'~S001R16 EE (Clmp Not Clsd, Slide Not Advd, Pin Not Retd, Still Opn, Still Ret) S001R16B#.O.A S001R16B#.I.## FB2[234].16'; 7505 '~S001R16 EE (Clmp Not Opnd, Slide Not Retd, Pin Not Advd, Still Clsd, Still Adv) S001R16B#.O.A S001R16B#.I.## FB2[234].17'; 7506 '~S001R16 EE (Clmp Not Clsd, Slide Not Advd, Pin Not Retd, Still Opn, Still Ret) S001R16B#.O.A S001R16B#.I.## FB2[234].18'; 7507 '~S001R16 EE (Clmp Not Opnd, Slide Not Retd, Pin Not Advd, Still Clsd, Still Adv) S001R16B#.O.A S001R16B#.I.## FB2[234].19'; 7508 '~S001R16 EE (Clmp Not Clsd, Slide Not Advd, Pin Not Retd, Still Opn, Still Ret) S001R16B#.O.A S001R16B#.I.## FB2[234].20'; 7509 '~S001R16 EE (Clmp Not Opnd, Slide Not Retd, Pin Not Advd, Still Clsd, Still Adv) S001R16B#.O.A S001R16B#.I.## FB2[234].21'; 7510 '~S001R16 EE (Clmp Not Clsd, Slide Not Advd, Pin Not Retd, Still Opn, Still Ret) S001R16B#.O.A S001R16B#.I.## FB2[234].22'; 7511 '~S001R16 EE (Clmp Not Opnd, Slide Not Retd, Pin Not Advd, Still Clsd, Still Adv) S001R16B#.O.A S001R16B#.I.## FB2[234].23'; 7512 '~S001R16 EE (Clmp Not Clsd, Slide Not Advd, Pin Not Retd, Still Opn, Still Ret) S001R16B#.O.A S001R16B#.I.## FB2[234].24'; 7513 '~S001R16 EE (Clmp Not Opnd, Slide Not Retd, Pin Not Advd, Still Clsd, Still Adv) S001R16B#.O.A S001R16B#.I.## FB2[234].25'; 7514 '~S001R16 EE (Clmp Not Clsd, Slide Not Advd, Pin Not Retd, Still Opn, Still Ret) S001R16B#.O.A S001R16B#.I.## FB2[234].26'; 7515 '~S001R16 EE (Clmp Not Opnd, Slide Not Retd, Pin Not Advd, Still Clsd, Still Adv) S001R16B#.O.A S001R16B#.I.## FB2[234].27'; 7516 '~S001R16 EE (Clmp Not Clsd, Slide Not Advd, Pin Not Retd, Still Opn, Still Ret) S001R16B#.O.A S001R16B#.I.## FB2[234].28'; 7517 '~S001R16 EE (Clmp Not Opnd, Slide Not Retd, Pin Not Advd, Still Clsd, Still Adv) S001R16B#.O.A S001R16B#.I.## FB2[234].29'; 7518 '~S001R16 EE (Clmp Not Clsd, Slide Not Advd, Pin Not Retd, Still Opn, Still Ret) S001R16B#.O.A S001R16B#.I.## FB2[234].30'; 7519 '~S001R16 EE (Clmp Not Opnd, Slide Not Retd, Pin Not Advd, Still Clsd, Still Adv) S001R16B#.O.A S001R16B#.I.## FB2[234].31'; 7520 '~S001R16 EE (Clmp Not Clsd, Slide Not Advd, Pin Not Retd, Still Opn, Still Ret) S001R16B#.O.A S001R16B#.I.## FB2[235].0'; 7521 '~S001R16 EE (Clmp Not Opnd, Slide Not Retd, Pin Not Advd, Still Clsd, Still Adv) S001R16B#.O.A S001R16B#.I.## FB2[235].1'; 7522 '~S001R16 EE (Clmp Not Clsd, Slide Not Advd, Pin Not Retd, Still Opn, Still Ret) S001R16B#.O.A S001R16B#.I.## FB2[235].2'; 7523 '~S001R16 EE (Clmp Not Opnd, Slide Not Retd, Pin Not Advd, Still Clsd, Still Adv) S001R16B#.O.A S001R16B#.I.## FB2[235].3'; 7524 '~S001R16 EE (Clmp Not Clsd, Slide Not Advd, Pin Not Retd, Still Opn, Still Ret) S001R16B#.O.A S001R16B#.I.## FB2[235].4'; 7525 '~S001R16 EE (Clmp Not Opnd, Slide Not Retd, Pin Not Advd, Still Clsd, Still Adv) S001R16B#.O.A S001R16B#.I.## FB2[235].5'; 7526 '~S001R16 EE (Clmp Not Clsd, Slide Not Advd, Pin Not Retd, Still Opn, Still Ret) S001R16B#.O.A S001R16B#.I.## FB2[235].6'; 7527 '~S001R16 EE (Clmp Not Opnd, Slide Not Retd, Pin Not Advd, Still Clsd, Still Adv) S001R16B#.O.A S001R16B#.I.## FB2[235].7'; 7528 '~S001R16 EE (Clmp Not Clsd, Slide Not Advd, Pin Not Retd, Still Opn, Still Ret) S001R16B#.O.A S001R16B#.I.## FB2[235].8'; 7529 '~S001R16 EE (Clmp Not Opnd, Slide Not Retd, Pin Not Advd, Still Clsd, Still Adv) S001R16B#.O.A S001R16B#.I.## FB2[235].9'; 7530 '~S001R16 EE (Clmp Not Clsd, Slide Not Advd, Pin Not Retd, Still Opn, Still Ret) S001R16B#.O.A S001R16B#.I.## FB2[235].10'; 7531 '~S001R16 EE (Clmp Not Opnd, Slide Not Retd, Pin Not Advd, Still Clsd, Still Adv) S001R16B#.O.A S001R16B#.I.## FB2[235].11'; 7532 '~S001R16 EE (Clmp Not Clsd, Slide Not Advd, Pin Not Retd, Still Opn, Still Ret) S001R16B#.O.A S001R16B#.I.## FB2[235].12'; 7533 '~S001R16 EE (Clmp Not Opnd, Slide Not Retd, Pin Not Advd, Still Clsd, Still Adv) S001R16B#.O.A S001R16B#.I.## FB2[235].13'; 7534 '~S001R16 EE (Clmp Not Clsd, Slide Not Advd, Pin Not Retd, Still Opn, Still Ret) S001R16B#.O.A S001R16B#.I.## FB2[235].14'; 7535 '~S001R16 EE (Clmp Not Opnd, Slide Not Retd, Pin Not Advd, Still Clsd, Still Adv) S001R16B#.O.A S001R16B#.I.## FB2[235].15'; 7536 '~S001R16 EE (Clmp Not Clsd, Slide Not Advd, Pin Not Retd, Still Opn, Still Ret) S001R16B#.O.A S001R16B#.I.## FB2[235].16'; 7537 '~S001R16 EE (Clmp Not Opnd, Slide Not Retd, Pin Not Advd, Still Clsd, Still Adv) S001R16B#.O.A S001R16B#.I.## FB2[235].17'; 7538 '~S001R16 EE (Clmp Not Clsd, Slide Not Advd, Pin Not Retd, Still Opn, Still Ret) S001R16B#.O.A S001R16B#.I.## FB2[235].18'; 7539 '~S001R16 EE (Clmp Not Opnd, Slide Not Retd, Pin Not Advd, Still Clsd, Still Adv) S001R16B#.O.A S001R16B#.I.## FB2[235].19'; 7540 '~S001R16 EE (Clmp Not Clsd, Slide Not Advd, Pin Not Retd, Still Opn, Still Ret) S001R16B#.O.A S001R16B#.I.## FB2[235].20'; 7541 '~S001R16 EE (Clmp Not Opnd, Slide Not Retd, Pin Not Advd, Still Clsd, Still Adv) S001R16B#.O.A S001R16B#.I.## FB2[235].21'; 7542 '~S001R16 EE (Clmp Not Clsd, Slide Not Advd, Pin Not Retd, Still Opn, Still Ret) S001R16B#.O.A S001R16B#.I.## FB2[235].22'; 7543 '~S001R16 EE (Clmp Not Opnd, Slide Not Retd, Pin Not Advd, Still Clsd, Still Adv) S001R16B#.O.A S001R16B#.I.## FB2[235].23'; 7544 '~S001R16 EE (Clmp Not Clsd, Slide Not Advd, Pin Not Retd, Still Opn, Still Ret) S001R16B#.O.A S001R16B#.I.## FB2[235].24'; 7545 '~S001R16 EE (Clmp Not Opnd, Slide Not Retd, Pin Not Advd, Still Clsd, Still Adv) S001R16B#.O.A S001R16B#.I.## FB2[235].25'; 7546 '~S001R16 EE (Clmp Not Clsd, Slide Not Advd, Pin Not Retd, Still Opn, Still Ret) S001R16B#.O.A S001R16B#.I.## FB2[235].26'; 7547 '~S001R16 EE (Clmp Not Opnd, Slide Not Retd, Pin Not Advd, Still Clsd, Still Adv) S001R16B#.O.A S001R16B#.I.## FB2[235].27'; 7548 '~S001R16 EE (Clmp Not Clsd, Slide Not Advd, Pin Not Retd, Still Opn, Still Ret) S001R16B#.O.A S001R16B#.I.## FB2[235].28'; 7549 '~S001R16 EE (Clmp Not Opnd, Slide Not Retd, Pin Not Advd, Still Clsd, Still Adv) S001R16B#.O.A S001R16B#.I.## FB2[235].29'; 7550 '~S001R16 EE (Clmp Not Clsd, Slide Not Advd, Pin Not Retd, Still Opn, Still Ret) S001R16B#.O.A S001R16B#.I.## FB2[235].30'; 7551 '~S001R16 EE (Clmp Not Opnd, Slide Not Retd, Pin Not Advd, Still Clsd, Still Adv) S001R16B#.O.A S001R16B#.I.## FB2[235].31'; 7552 '~Spare FB2[236].0'; 7553 '~Spare FB2[236].1'; 7554 '~Spare FB2[236].2'; 7555 '~Spare FB2[236].3'; 7556 '~Spare FB2[236].4'; 7557 '~Spare FB2[236].5'; 7558 '~Spare FB2[236].6'; 7559 '~Spare FB2[236].7'; 7560 '~Spare FB2[236].8'; 7561 '~Spare FB2[236].9'; 7562 '~Spare FB2[236].10'; 7563 '~Spare FB2[236].11'; 7564 '~Spare FB2[236].12'; 7565 '~Spare FB2[236].13'; 7566 '~Spare FB2[236].14'; 7567 '~Spare FB2[236].15'; 7568 '~Spare FB2[236].16'; 7569 '~Spare FB2[236].17'; 7570 '~Spare FB2[236].18'; 7571 '~Spare FB2[236].19'; 7572 '~Spare FB2[236].20'; 7573 '~Spare FB2[236].21'; 7574 '~Spare FB2[236].22'; 7575 '~Spare FB2[236].23'; 7576 '~Spare FB2[236].24'; 7577 '~Spare FB2[236].25'; 7578 '~Spare FB2[236].26'; 7579 '~Spare FB2[236].27'; 7580 '~Spare FB2[236].28'; 7581 '~Spare FB2[236].29'; 7582 '~Spare FB2[236].30'; 7583 '~Spare FB2[236].31'; 7584 '~Spare FB2[237].0'; 7585 '~Spare FB2[237].1'; 7586 '~Spare FB2[237].2'; 7587 '~Spare FB2[237].3'; 7588 '~Spare FB2[237].4'; 7589 '~Spare FB2[237].5'; 7590 '~Spare FB2[237].6'; 7591 '~Spare FB2[237].7'; 7592 '~Spare FB2[237].8'; 7593 '~Spare FB2[237].9'; 7594 '~Spare FB2[237].10'; 7595 '~Spare FB2[237].11'; 7596 '~Spare FB2[237].12'; 7597 '~Spare FB2[237].13'; 7598 '~Spare FB2[237].14'; 7599 '~Spare FB2[237].15'; 7600 '~Spare FB2[237].16'; 7601 '~Spare FB2[237].17'; 7602 '~Spare FB2[237].18'; 7603 '~Spare FB2[237].19'; 7604 '~Spare FB2[237].20'; 7605 '~Spare FB2[237].21'; 7606 '~Spare FB2[237].22'; 7607 '~Spare FB2[237].23'; 7608 '~Spare FB2[237].24'; 7609 '~Spare FB2[237].25'; 7610 '~Spare FB2[237].26'; 7611 '~Spare FB2[237].27'; 7612 '~Spare FB2[237].28'; 7613 '~Spare FB2[237].29'; 7614 '~Spare FB2[237].30'; 7615 '~Spare FB2[237].31'; 7616 '~Spare FB2[238].0'; 7617 '~Spare FB2[238].1'; 7618 '~Spare FB2[238].2'; 7619 '~Spare FB2[238].3'; 7620 '~Spare FB2[238].4'; 7621 '~Spare FB2[238].5'; 7622 '~Spare FB2[238].6'; 7623 '~Spare FB2[238].7'; 7624 '~Spare FB2[238].8'; 7625 '~Spare FB2[238].9'; 7626 '~Spare FB2[238].10'; 7627 '~Spare FB2[238].11'; 7628 '~Spare FB2[238].12'; 7629 '~Spare FB2[238].13'; 7630 '~Spare FB2[238].14'; 7631 '~Spare FB2[238].15'; 7632 '~Spare FB2[238].16'; 7633 '~Spare FB2[238].17'; 7634 '~Spare FB2[238].18'; 7635 '~Spare FB2[238].19'; 7636 '~Spare FB2[238].20'; 7637 '~Spare FB2[238].21'; 7638 '~Spare FB2[238].22'; 7639 '~Spare FB2[238].23'; 7640 '~Spare FB2[238].24'; 7641 '~Spare FB2[238].25'; 7642 '~Spare FB2[238].26'; 7643 '~Spare FB2[238].27'; 7644 '~Spare FB2[238].28'; 7645 '~Spare FB2[238].29'; 7646 '~Spare FB2[238].30'; 7647 '~Spare FB2[238].31'; 7648 '~S001R16 (Peripheral Tool 1) Vlv/Otpt 1 Failed S001R16F#B#.O.# (Cls Clmps, Adv Slide, Ret Pins) FB2[239].0'; 7649 '~S001R16 (Peripheral Tool 1) Vlv/Otpt 1 Failed S001R16F#B#.O.# (Opn Clmps, Ret Slide, Adv Pins) FB2[239].1'; 7650 '~S001R16 (Peripheral Tool 1) Vlv/Otpt 2 Failed S001R16F#B#.O.# (Cls Clmps, Adv Slide, Ret Pins) FB2[239].2'; 7651 '~S001R16 (Peripheral Tool 1) Vlv/Otpt 2 Failed S001R16F#B#.O.# (Opn Clmps, Ret Slide, Adv Pins) FB2[239].3'; 7652 '~S001R16 (Peripheral Tool 1) Vlv/Otpt 3 Failed S001R16F#B#.O.# (Cls Clmps, Adv Slide, Ret Pins) FB2[239].4'; 7653 '~S001R16 (Peripheral Tool 1) Vlv/Otpt 3 Failed S001R16F#B#.O.# (Opn Clmps, Ret Slide, Adv Pins) FB2[239].5'; 7654 '~S001R16 (Peripheral Tool 1) Vlv/Otpt 4 Failed S001R16F#B#.O.# (Cls Clmps, Adv Slide, Ret Pins) FB2[239].6'; 7655 '~S001R16 (Peripheral Tool 1) Vlv/Otpt 4 Failed S001R16F#B#.O.# (Opn Clmps, Ret Slide, Adv Pins) FB2[239].7'; 7656 '~U-#### (Clmp Not Clsd, Slide Not Advd, Pin Not Retd, Still Opnd, Still Retd) S001R16F#.B#.O.# FB2[239].8'; 7657 '~U-#### (Clmp Not Opnd, Slide Not Retd, Pin Not Advd, Still Clsd, Still Advd) S001R16F#.B#.O.# FB2[239].9'; 7658 '~U-#### (Clmp Not Clsd, Slide Not Advd, Pin Not Retd, Still Opnd, Still Retd) S001R16F#.B#.O.# FB2[239].10'; 7659 '~U-#### (Clmp Not Opnd, Slide Not Retd, Pin Not Advd, Still Clsd, Still Advd) S001R16F#.B#.O.# FB2[239].11'; 7660 '~U-#### (Clmp Not Clsd, Slide Not Advd, Pin Not Retd, Still Opnd, Still Retd) S001R16F#.B#.O.# FB2[239].12'; 7661 '~U-#### (Clmp Not Opnd, Slide Not Retd, Pin Not Advd, Still Clsd, Still Advd) S001R16F#.B#.O.# FB2[239].13'; 7662 '~U-#### (Clmp Not Clsd, Slide Not Advd, Pin Not Retd, Still Opnd, Still Retd) S001R16F#.B#.O.# FB2[239].14'; 7663 '~U-#### (Clmp Not Opnd, Slide Not Retd, Pin Not Advd, Still Clsd, Still Advd) S001R16F#.B#.O.# FB2[239].15'; 7664 '~S001R16 (Peripheral Tool 2) Vlv/Otpt 1 Failed S001R16F#B#.O.# (Cls Clmps, Adv Slide, Ret Pins) FB2[239].16'; 7665 '~S001R16 (Peripheral Tool 2) Vlv/Otpt 1 Failed S001R16F#B#.O.# (Opn Clmps, Ret Slide, Adv Pins) FB2[239].17'; 7666 '~S001R16 (Peripheral Tool 2) Vlv/Otpt 2 Failed S001R16F#B#.O.# (Cls Clmps, Adv Slide, Ret Pins) FB2[239].18'; 7667 '~S001R16 (Peripheral Tool 2) Vlv/Otpt 2 Failed S001R16F#B#.O.# (Opn Clmps, Ret Slide, Adv Pins) FB2[239].19'; 7668 '~S001R16 (Peripheral Tool 2) Vlv/Otpt 3 Failed S001R16F#B#.O.# (Cls Clmps, Adv Slide, Ret Pins) FB2[239].20'; 7669 '~S001R16 (Peripheral Tool 2) Vlv/Otpt 3 Failed S001R16F#B#.O.# (Opn Clmps, Ret Slide, Adv Pins) FB2[239].21'; 7670 '~S001R16 (Peripheral Tool 2) Vlv/Otpt 4 Failed S001R16F#B#.O.# (Cls Clmps, Adv Slide, Ret Pins) FB2[239].22'; 7671 '~S001R16 (Peripheral Tool 2) Vlv/Otpt 4 Failed S001R16F#B#.O.# (Opn Clmps, Ret Slide, Adv Pins) FB2[239].23'; 7672 '~U-#### (Clmp Not Clsd, Slide Not Advd, Pin Not Retd, Still Opnd, Still Retd) S001R16F#.B#.O.# FB2[239].24'; 7673 '~U-#### (Clmp Not Opnd, Slide Not Retd, Pin Not Advd, Still Clsd, Still Advd) S001R16F#.B#.O.# FB2[239].25'; 7674 '~U-#### (Clmp Not Clsd, Slide Not Advd, Pin Not Retd, Still Opnd, Still Retd) S001R16F#.B#.O.# FB2[239].26'; 7675 '~U-#### (Clmp Not Opnd, Slide Not Retd, Pin Not Advd, Still Clsd, Still Advd) S001R16F#.B#.O.# FB2[239].27'; 7676 '~U-#### (Clmp Not Clsd, Slide Not Advd, Pin Not Retd, Still Opnd, Still Retd) S001R16F#.B#.O.# FB2[239].28'; 7677 '~U-#### (Clmp Not Opnd, Slide Not Retd, Pin Not Advd, Still Clsd, Still Advd) S001R16F#.B#.O.# FB2[239].29'; 7678 '~U-#### (Clmp Not Clsd, Slide Not Advd, Pin Not Retd, Still Opnd, Still Retd) S001R16F#.B#.O.# FB2[239].30'; 7679 '~U-#### (Clmp Not Opnd, Slide Not Retd, Pin Not Advd, Still Clsd, Still Advd) S001R16F#.B#.O.# FB2[239].31'; 7680 '~Spare FB2[240].0'; 7681 '~Spare FB2[240].1'; 7682 '~Spare FB2[240].2'; 7683 '~Spare FB2[240].3'; 7684 '~Spare FB2[240].4'; 7685 '~Spare FB2[240].5'; 7686 '~Spare FB2[240].6'; 7687 '~Spare FB2[240].7'; 7688 '~Spare FB2[240].8'; 7689 '~Spare FB2[240].9'; 7690 '~Spare FB2[240].10'; 7691 '~Spare FB2[240].11'; 7692 '~Spare FB2[240].12'; 7693 '~Spare FB2[240].13'; 7694 '~Spare FB2[240].14'; 7695 '~Spare FB2[240].15'; 7696 '~Spare FB2[240].16'; 7697 '~Spare FB2[240].17'; 7698 '~Spare FB2[240].18'; 7699 '~Spare FB2[240].19'; 7700 '~Spare FB2[240].20'; 7701 '~Spare FB2[240].21'; 7702 '~Spare FB2[240].22'; 7703 '~Spare FB2[240].23'; 7704 '~Spare FB2[240].24'; 7705 '~Spare FB2[240].25'; 7706 '~Spare FB2[240].26'; 7707 '~Spare FB2[240].27'; 7708 '~Spare FB2[240].28'; 7709 '~Spare FB2[240].29'; 7710 '~Spare FB2[240].30'; 7711 '~Spare FB2[240].31'; 7712 '~Spare FB2[241].0'; 7713 '~Spare FB2[241].1'; 7714 '~Spare FB2[241].2'; 7715 '~Spare FB2[241].3'; 7716 '~Spare FB2[241].4'; 7717 '~Spare FB2[241].5'; 7718 '~Spare FB2[241].6'; 7719 '~Spare FB2[241].7'; 7720 '~Spare FB2[241].8'; 7721 '~Spare FB2[241].9'; 7722 '~Spare FB2[241].10'; 7723 '~Spare FB2[241].11'; 7724 '~Spare FB2[241].12'; 7725 '~Spare FB2[241].13'; 7726 '~Spare FB2[241].14'; 7727 '~Spare FB2[241].15'; 7728 '~Spare FB2[241].16'; 7729 '~Spare FB2[241].17'; 7730 '~Spare FB2[241].18'; 7731 '~Spare FB2[241].19'; 7732 '~Spare FB2[241].20'; 7733 '~Spare FB2[241].21'; 7734 '~Spare FB2[241].22'; 7735 '~Spare FB2[241].23'; 7736 '~Spare FB2[241].24'; 7737 '~Spare FB2[241].25'; 7738 '~Spare FB2[241].26'; 7739 '~Spare FB2[241].27'; 7740 '~Spare FB2[241].28'; 7741 '~Spare FB2[241].29'; 7742 '~Spare FB2[241].30'; 7743 '~Spare FB2[241].31'; 7744 '~Spare FB2[242].0'; 7745 '~Spare FB2[242].1'; 7746 '~Spare FB2[242].2'; 7747 '~Spare FB2[242].3'; 7748 '~Spare FB2[242].4'; 7749 '~Spare FB2[242].5'; 7750 '~Spare FB2[242].6'; 7751 '~Spare FB2[242].7'; 7752 '~Spare FB2[242].8'; 7753 '~Spare FB2[242].9'; 7754 '~Spare FB2[242].10'; 7755 '~Spare FB2[242].11'; 7756 '~Spare FB2[242].12'; 7757 '~Spare FB2[242].13'; 7758 '~Spare FB2[242].14'; 7759 '~Spare FB2[242].15'; 7760 '~Spare FB2[242].16'; 7761 '~Spare FB2[242].17'; 7762 '~Spare FB2[242].18'; 7763 '~Spare FB2[242].19'; 7764 '~Spare FB2[242].20'; 7765 '~Spare FB2[242].21'; 7766 '~Spare FB2[242].22'; 7767 '~Spare FB2[242].23'; 7768 '~Spare FB2[242].24'; 7769 '~Spare FB2[242].25'; 7770 '~Spare FB2[242].26'; 7771 '~Spare FB2[242].27'; 7772 '~Spare FB2[242].28'; 7773 '~Spare FB2[242].29'; 7774 '~Spare FB2[242].30'; 7775 '~Spare FB2[242].31'; 7776 '~Spare FB2[243].0'; 7777 '~Spare FB2[243].1'; 7778 '~Spare FB2[243].2'; 7779 '~Spare FB2[243].3'; 7780 '~Spare FB2[243].4'; 7781 '~Spare FB2[243].5'; 7782 '~Spare FB2[243].6'; 7783 '~Spare FB2[243].7'; 7784 '~Spare FB2[243].8'; 7785 '~Spare FB2[243].9'; 7786 '~Spare FB2[243].10'; 7787 '~Spare FB2[243].11'; 7788 '~Spare FB2[243].12'; 7789 '~Spare FB2[243].13'; 7790 '~Spare FB2[243].14'; 7791 '~Spare FB2[243].15'; 7792 '~Spare FB2[243].16'; 7793 '~Spare FB2[243].17'; 7794 '~Spare FB2[243].18'; 7795 '~Spare FB2[243].19'; 7796 '~Spare FB2[243].20'; 7797 '~Spare FB2[243].21'; 7798 '~Spare FB2[243].22'; 7799 '~Spare FB2[243].23'; 7800 '~Spare FB2[243].24'; 7801 '~Spare FB2[243].25'; 7802 '~Spare FB2[243].26'; 7803 '~Spare FB2[243].27'; 7804 '~Spare FB2[243].28'; 7805 '~Spare FB2[243].29'; 7806 '~Spare FB2[243].30'; 7807 '~Spare FB2[243].31'; 7808 '~S001R09CN.I.RbtCtrlFlt - Control Fault FB2[244].0'; 7809 '~S001R09CN.I.CollDetect - Collision Detect FB2[244].1'; 7810 '~S001R09CN.Ix.RbtPromptBox - View Prompt Box at Teach Pendant FB2[244].2'; 7811 '~Spare FB2[244].3'; 7812 '~Spare FB2[244].4'; 7813 '~Spare FB2[244].5'; 7814 '~Spare FB2[244].6'; 7815 '~Spare FB2[244].7'; 7816 '~Spare FB2[244].8'; 7817 '~Spare FB2[244].9'; 7818 '~Spare FB2[244].10'; 7819 '~S001R09CN.I.Wc1WldFlt -Weld Controller 1 Weld Fault FB2[244].11'; 7820 '~S001R09CN.I.Wc1Flt - Weld Timer Flt - Depress Man Weld To Continue FB2[244].12'; 7821 '~S001R09CN.I.Wc1SGunFlt - Weld Controller 1 Servo Gun Fault FB2[244].13'; 7822 '~S001R09CN.I.Wc1SGunMtrTempFlt - Cntrl 1 Servo Gun Motor Over Temp FB2[244].14'; 7823 '~S001R09CN.I.Td1MtrFlt - Tip Dress 1 Motor Fault FB2[244].15'; 7824 '~S001R09CN.I.WC1XfmrTempFlt - Weld Cntrl 1 Transformer Over Temp FB2[244].16'; 7825 '~S001R09CN.I.AutoTipChng1Flt - Auto Tip Changer 1 Fault FB2[244].17'; 7826 '~S001R09CN.I.Slr1NotReady - Seal Controller 1 Not Ready FB2[244].18'; 7827 '~S001R09CN.I.Slr1MajorFlt - Seal Controller 1 Major Fault FB2[244].19'; 7828 '~S001R09CN.I.Slr1VolNotOk - Seal Controller 1 Volume Not Ok Fault FB2[244].20'; 7829 '~S001R09CN.I.Slr1PurgeFlt - Seal Controller 1 Purge Fault FB2[244].21'; 7830 '~S001R09CN.I.Slr1DoserNot Filled - Seal Cntrl 1 Doser Not Filled FB2[244].22'; 7831 '~S001R09CN.I.Slr1No2ClnMxr - Seal Cntrl1 No 2C In Mixer Fault FB2[244].23'; 7832 '~S001R09CN.I.Slr1NzlBroken - Seal Controller 1 Nozzle Broken Fault FB2[244].24'; 7833 '~S001R09CN.I.Slr1NozzleChgReq - Seal Cntrl1 Nozzle Change Reqd FB2[244].25'; 7834 '~S001R09CN.I.Slr1CycleInterrupted - Seal Cntrl1 Cycle Interrupted FB2[244].26'; 7835 '~S001R09CN.I.Stdw1Flt - Stud Weld 1 Weld Fault FB2[244].27'; 7836 '~S001R09CN.I.Stdw1DlyExcdd - Stud Weld 1 Time Delay Exceeded Flt FB2[244].28'; 7837 '~S001R09CN.I.Stdw1Maint Reqd - Stud Weld 1 Maintenance Required FB2[244].29'; 7838 '~S001R09CN.I.Stdw1Reject - Stud Weld 1 art Reject Fault FB2[244].30'; 7839 '~S001R09CN.I.Rvt1Flt - Rivet Controller 1 Fault FB2[244].31'; 7840 '~S001R09CN.I.Rvt1DlyExcdd - Rivet Cntrl 1 Time Delay Exceeded Flt FB2[245].0'; 7841 '~S001R09CN.I.AutoPulledTipByp1 - Auto Pulled Tip Bypass 1 FB2[245].1'; 7842 '~S001R09CN.I.StdWld1EquipmentFlt - Stud Weld 1 Equipment Fault FB2[245].2'; 7843 '~S001R09CN.I.StdWld1BrcktNotPresent - Stud Weld 1 Bracket Not Pres FB2[245].3'; 7844 '~S001R09CN.I.PierceFlt - Pierce Fault FB2[245].4'; 7845 '~S001R09CN.I.NoVisionMeasErr - Vision System Measurement Error FB2[245].5'; 7846 '~S001R09CN.I.VisionSysCalErr - Vision System Calibration Fault FB2[245].6'; 7847 '~S001R09CN.I.VisionSysErr - Vision System Error FB2[245].7'; 7848 '~S001R09CN.I.RackOutOfTolerance - Vision Sys Rack Out Of Tolerance FB2[245].8'; 7849 '~S001R09CN.Ix.TorqFlt - Torque Not Ok FB2[245].9'; 7850 '~S001R09CN.Ix.MwFlt - Mig Weld Controller Fault FB2[245].10'; 7851 '~S001R09CN.Ix.MwWireStuckFlt - Mig Welder Wire Stuck FB2[245].11'; 7852 '~S001R09CN.Ix.MwWldFlt - Mig Welder Bad Bronze Weld Indicator Flt FB2[245].12'; 7853 '~S001R09CN.I.O.TipChngReqd1 - Weld Cntrl 1 Tip Change Required FB2[245].13'; 7854 '~S001R09CN.I.M.NutDetectFlt1 - Nut Welder 1 Nut Detection Fault FB2[245].14'; 7855 '~S001R09CN.I.M.NutProjFlt1 - Nut Welder 1 Weld Not In Tolerance FB2[245].15'; 7856 '~S001R09CN.M.WrongRivetAtNose - Remove Wrong Rivet At Nose FB2[245].16'; 7857 '~S001R09CN.Ix.MwWldLimitErr - Mig Welder CurrentVoltage Out of Tolerance FB2[245].17'; 7858 '~S001R09CN.Ix.MigRdy Mig Welder Not Ready FB2[245].18'; 7859 '~Spare FB2[245].19'; 7860 '~Spare FB2[245].20'; 7861 '~S001R09CN.I.Wc2WldFlt -Weld Controller 2 Weld Fault FB2[245].21'; 7862 '~S001R09CN.I.Wc2Flt - Weld Timer Flt - Depress Man Weld To Continue FB2[245].22'; 7863 '~S001R09CN.I.Wc2SGunFlt - Weld Controller 2 Servo Gun Fault FB2[245].23'; 7864 '~S001R09CN.I.Wc2SGunMtrTempFlt - Cntrl 2 Servo Gun Motor Over Temp FB2[245].24'; 7865 '~S001R09CN.I.Td2MtrFlt - Tip Dress 2 Motor Fault FB2[245].25'; 7866 '~S001R09CN.I.WC2XfmrTempFlt - Weld Cntrl 2 Transformer Over Temp FB2[245].26'; 7867 '~S001R09CN.I.AutoTipChng2Flt - Auto Tip Changer 2 Fault FB2[245].27'; 7868 '~S001R09CN.I.Slr2NotReady - Seal Controller 2 Not Ready FB2[245].28'; 7869 '~S001R09CN.I.Slr2MajorFlt - Seal Controller 2 Major Fault FB2[245].29'; 7870 '~S001R09CN.I.Slr2VolNotOk - Seal Controller 2 Volume Not Ok Fault FB2[245].30'; 7871 '~S001R09CN.I.Slr2PurgeFlt - Seal Controller 2 Purge Fault FB2[245].31'; 7872 '~S001R09CN.I.Slr2DoserNot Filled - Seal Cntrl 2 Doser Not Filled FB2[246].0'; 7873 '~S001R09CN.I.Slr2No2ClnMxr - Seal Cntrl2 No 2C In Mixer Fault FB2[246].1'; 7874 '~S001R09CN.I.Slr2NzlBroken - Seal Controller 2 Nozzle Broken Fault FB2[246].2'; 7875 '~S001R09CN.I.Slr2NozzleChgReq - Seal Cntrl2 Nozzle Change Reqd FB2[246].3'; 7876 '~S001R09CN.I.Slr2CycleInterrupted - Seal Cntrl2 Cycle Interrupted FB2[246].4'; 7877 '~S001R09CN.I.Stdw2Flt - Stud Weld 2 Weld Fault FB2[246].5'; 7878 '~S001R09CN.I.Stdw2DlyExcdd - Stud Weld 2 Time Delay Exceeded Flt FB2[246].6'; 7879 '~S001R09CN.I.Stdw2Maint Reqd - Stud Weld 2 Maintenance Required FB2[246].7'; 7880 '~S001R09CN.I.Stdw2Reject - Stud Weld 2 art Reject Fault FB2[246].8'; 7881 '~S001R09CN.I.Rvt2Flt - Rivet Controller 2 Fault FB2[246].9'; 7882 '~S001R09CN.I.Rvt2DlyExcdd - Rivet Cntrl 2 Time Delay Exceeded Flt FB2[246].10'; 7883 '~S001R09CN.I.AutoPulledTipByp2 - Auto Pulled Tip Bypass 2 FB2[246].11'; 7884 '~S001R09CN.I.StdWld2EquipmentFlt - Stud Weld 2 Equipment Fault FB2[246].12'; 7885 '~S001R09CN.I.StdWld2BrcktNotPresent - Stud Weld 2 Bracket Not Pres FB2[246].13'; 7886 '~S001R09CN.Ix.LsrWldMntrFlt - Seam Geometry/Laser Weld Monitor Flt FB2[246].14'; 7887 '~S001R09CN.Ix.LsrHeadFlt - Laser Head Fault FB2[246].15'; 7888 '~S001R09CN.Ix.LsrGlsFlt - Glass Fault FB2[246].16'; 7889 '~S001R09CN.Ix.LsrWhlFlt - Pressure Wheel Not In Range Fault FB2[246].17'; 7890 '~S001R09CN.Ix.LsrGeoFlt - Seam Geometry/Laser Bad Process Geo Flt FB2[246].18'; 7891 '~S001R09CN.Ix.LsrHdCollFlt - Laser Head Collision Fault FB2[246].19'; 7892 '~S001R09CN.Ix.LsrHdSysFlt - Laser Head System Fault FB2[246].20'; 7893 '~S001R09CN.Ix.LsrHdFar - Laser Head Far Fault FB2[246].21'; 7894 '~S001R09CN.Ix.LsrHdSftCollFlt - Laser Head Software Collision Flt FB2[246].22'; 7895 '~S001R09CN.I.O.TipChngReqd2 - Weld Cntrl 2 Tip Change Required FB2[246].23'; 7896 '~S001R09CN.I.M.NutDetectFlt2 - Nut Welder 2 Nut Detection Fault FB2[246].24'; 7897 '~S001R09CN.I.M.NutProjFlt2 - Nut Welder 2 Weld Not In Tolerance FB2[246].25'; 7898 '~S001R09CN.I.TCWrongToolInStand - Tool Changer Wrong Tool In Stand FB2[246].26'; 7899 '~Spare FB2[246].27'; 7900 '~Spare FB2[246].28'; 7901 '~Spare FB2[246].29'; 7902 '~Spare FB2[246].30'; 7903 '~Spare FB2[246].31'; 7904 '~S001R09CN.I.VisionCommOK - Vision System Comm Fault FB2[247].0'; 7905 '~S001R09CN.I.OutOfTolerance - Vision System Out Of Tolerance FB2[247].1'; 7906 '~S001R09CN.I.MeasureReject - Vision System Measure Reject FB2[247].2'; 7907 '~S001R09CN.I.VisionSysCalibrationFlt - Vision System Calibration Flt FB2[247].3'; 7908 '~S001R09CN.I.VisionSysFlt - Vision System Flt FB2[247].4'; 7909 '~Spare FB2[247].5'; 7910 '~Spare FB2[247].6'; 7911 '~Spare FB2[247].7'; 7912 '~Spare FB2[247].8'; 7913 '~Spare FB2[247].9'; 7914 '~Spare FB2[247].10'; 7915 '~Spare FB2[247].11'; 7916 '~Spare FB2[247].12'; 7917 '~Spare FB2[247].13'; 7918 '~Spare FB2[247].14'; 7919 '~Spare FB2[247].15'; 7920 '~Spare FB2[247].16'; 7921 '~Spare FB2[247].17'; 7922 '~S001R09CN.M.InteruptCyc - Laser Cyc Interupt Cut Wire And Reject Car FB2[247].18'; 7923 '~S001R09CN.M.SuspectPart Inspect Vehicle And Accept Or Reject FB2[247].19'; 7924 '~S001R09 Power Meter High Power Fault Detected FB2[247].20'; 7925 '~S001R09 Power Meter Low Power Fault Detected FB2[247].21'; 7926 '~Spare FB2[247].22'; 7927 '~Spare FB2[247].23'; 7928 '~Spare FB2[247].24'; 7929 '~Spare FB2[247].25'; 7930 '~Spare FB2[247].26'; 7931 '~Spare FB2[247].27'; 7932 '~Spare FB2[247].28'; 7933 '~Spare FB2[247].29'; 7934 '~Spare FB2[247].30'; 7935 '~Spare FB2[247].31'; 7936 '~Spare FB2[248].0'; 7937 '~Spare FB2[248].1'; 7938 '~Spare FB2[248].2'; 7939 '~Spare FB2[248].3'; 7940 '~Spare FB2[248].4'; 7941 '~Spare FB2[248].5'; 7942 '~Spare FB2[248].6'; 7943 '~Spare FB2[248].7'; 7944 '~Spare FB2[248].8'; 7945 '~Spare FB2[248].9'; 7946 '~Spare FB2[248].10'; 7947 '~Spare FB2[248].11'; 7948 '~Spare FB2[248].12'; 7949 '~Spare FB2[248].13'; 7950 '~Spare FB2[248].14'; 7951 '~Spare FB2[248].15'; 7952 '~Spare FB2[248].16'; 7953 '~Spare FB2[248].17'; 7954 '~Spare FB2[248].18'; 7955 '~Spare FB2[248].19'; 7956 '~Spare FB2[248].20'; 7957 '~Spare FB2[248].21'; 7958 '~Spare FB2[248].22'; 7959 '~Spare FB2[248].23'; 7960 '~Spare FB2[248].24'; 7961 '~Spare FB2[248].25'; 7962 '~Spare FB2[248].26'; 7963 '~Spare FB2[248].27'; 7964 '~Spare FB2[248].28'; 7965 '~Spare FB2[248].29'; 7966 '~Spare FB2[248].30'; 7967 '~Spare FB2[248].31'; 7968 '~Spare FB2[249].0'; 7969 '~Spare FB2[249].1'; 7970 '~Spare FB2[249].2'; 7971 '~Spare FB2[249].3'; 7972 '~Spare FB2[249].4'; 7973 '~Spare FB2[249].5'; 7974 '~Spare FB2[249].6'; 7975 '~Spare FB2[249].7'; 7976 '~Spare FB2[249].8'; 7977 '~Spare FB2[249].9'; 7978 '~Spare FB2[249].10'; 7979 '~Spare FB2[249].11'; 7980 '~Spare FB2[249].12'; 7981 '~Spare FB2[249].13'; 7982 '~Spare FB2[249].14'; 7983 '~Spare FB2[249].15'; 7984 '~Spare FB2[249].16'; 7985 '~Spare FB2[249].17'; 7986 '~Spare FB2[249].18'; 7987 '~Spare FB2[249].19'; 7988 '~Spare FB2[249].20'; 7989 '~Spare FB2[249].21'; 7990 '~Spare FB2[249].22'; 7991 '~Spare FB2[249].23'; 7992 '~Spare FB2[249].24'; 7993 '~Spare FB2[249].25'; 7994 '~Spare FB2[249].26'; 7995 '~Spare FB2[249].27'; 7996 '~Spare FB2[249].28'; 7997 '~Spare FB2[249].29'; 7998 '~Spare FB2[249].30'; 7999 '~Spare FB2[249].31'; 8000 '~Spare FB2[250].0'; 8001 '~Spare FB2[250].1'; 8002 '~Spare FB2[250].2'; 8003 '~Spare FB2[250].3'; 8004 '~Spare FB2[250].4'; 8005 '~Spare FB2[250].5'; 8006 '~Spare FB2[250].6'; 8007 '~Spare FB2[250].7'; 8008 '~Spare FB2[250].8'; 8009 '~Spare FB2[250].9'; 8010 '~Spare FB2[250].10'; 8011 '~Spare FB2[250].11'; 8012 '~Spare FB2[250].12'; 8013 '~Spare FB2[250].13'; 8014 '~Spare FB2[250].14'; 8015 '~Spare FB2[250].15'; 8016 '~Spare FB2[250].16'; 8017 '~Spare FB2[250].17'; 8018 '~Spare FB2[250].18'; 8019 '~Spare FB2[250].19'; 8020 '~Spare FB2[250].20'; 8021 '~Spare FB2[250].21'; 8022 '~Spare FB2[250].22'; 8023 '~Spare FB2[250].23'; 8024 '~Spare FB2[250].24'; 8025 '~Spare FB2[250].25'; 8026 '~Spare FB2[250].26'; 8027 '~Spare FB2[250].27'; 8028 '~Spare FB2[250].28'; 8029 '~Spare FB2[250].29'; 8030 '~Spare FB2[250].30'; 8031 '~Spare FB2[250].31'; 8032 '~Spare FB2[251].0'; 8033 '~Spare FB2[251].1'; 8034 '~Spare FB2[251].2'; 8035 '~Spare FB2[251].3'; 8036 '~Spare FB2[251].4'; 8037 '~Spare FB2[251].5'; 8038 '~Spare FB2[251].6'; 8039 '~Spare FB2[251].7'; 8040 '~Spare FB2[251].8'; 8041 '~Spare FB2[251].9'; 8042 '~Spare FB2[251].10'; 8043 '~Spare FB2[251].11'; 8044 '~Spare FB2[251].12'; 8045 '~Spare FB2[251].13'; 8046 '~Spare FB2[251].14'; 8047 '~Spare FB2[251].15'; 8048 '~Spare FB2[251].16'; 8049 '~Spare FB2[251].17'; 8050 '~Spare FB2[251].18'; 8051 '~Spare FB2[251].19'; 8052 '~Spare FB2[251].20'; 8053 '~Spare FB2[251].21'; 8054 '~Spare FB2[251].22'; 8055 '~Spare FB2[251].23'; 8056 '~Spare FB2[251].24'; 8057 '~Spare FB2[251].25'; 8058 '~Spare FB2[251].26'; 8059 '~Spare FB2[251].27'; 8060 '~Spare FB2[251].28'; 8061 '~Spare FB2[251].29'; 8062 '~Spare FB2[251].30'; 8063 '~Spare FB2[251].31'; 8064 '~S001R10CN.I.RbtCtrlFlt - Control Fault FB2[252].0'; 8065 '~S001R10CN.I.CollDetect - Collision Detect FB2[252].1'; 8066 '~S001R10CN.Ix.RbtPromptBox - View Prompt Box at Teach Pendant FB2[252].2'; 8067 '~Spare FB2[252].3'; 8068 '~Spare FB2[252].4'; 8069 '~Spare FB2[252].5'; 8070 '~Spare FB2[252].6'; 8071 '~Spare FB2[252].7'; 8072 '~Spare FB2[252].8'; 8073 '~Spare FB2[252].9'; 8074 '~Spare FB2[252].10'; 8075 '~S001R10CN.I.Wc1WldFlt -Weld Controller 1 Weld Fault FB2[252].11'; 8076 '~S001R10CN.I.Wc1Flt - Weld Timer Flt - Depress Man Weld To Continue FB2[252].12'; 8077 '~S001R10CN.I.Wc1SGunFlt - Weld Controller 1 Servo Gun Fault FB2[252].13'; 8078 '~S001R10CN.I.Wc1SGunMtrTempFlt - Cntrl 1 Servo Gun Motor Over Temp FB2[252].14'; 8079 '~S001R10CN.I.Td1MtrFlt - Tip Dress 1 Motor Fault FB2[252].15'; 8080 '~S001R10CN.I.WC1XfmrTempFlt - Weld Cntrl 1 Transformer Over Temp FB2[252].16'; 8081 '~S001R10CN.I.AutoTipChng1Flt - Auto Tip Changer 1 Fault FB2[252].17'; 8082 '~S001R10CN.I.Slr1NotReady - Seal Controller 1 Not Ready FB2[252].18'; 8083 '~S001R10CN.I.Slr1MajorFlt - Seal Controller 1 Major Fault FB2[252].19'; 8084 '~S001R10CN.I.Slr1VolNotOk - Seal Controller 1 Volume Not Ok Fault FB2[252].20'; 8085 '~S001R10CN.I.Slr1PurgeFlt - Seal Controller 1 Purge Fault FB2[252].21'; 8086 '~S001R10CN.I.Slr1DoserNot Filled - Seal Cntrl 1 Doser Not Filled FB2[252].22'; 8087 '~S001R10CN.I.Slr1No2ClnMxr - Seal Cntrl1 No 2C In Mixer Fault FB2[252].23'; 8088 '~S001R10CN.I.Slr1NzlBroken - Seal Controller 1 Nozzle Broken Fault FB2[252].24'; 8089 '~S001R10CN.I.Slr1NozzleChgReq - Seal Cntrl1 Nozzle Change Reqd FB2[252].25'; 8090 '~S001R10CN.I.Slr1CycleInterrupted - Seal Cntrl1 Cycle Interrupted FB2[252].26'; 8091 '~S001R10CN.I.Stdw1Flt - Stud Weld 1 Weld Fault FB2[252].27'; 8092 '~S001R10CN.I.Stdw1DlyExcdd - Stud Weld 1 Time Delay Exceeded Flt FB2[252].28'; 8093 '~S001R10CN.I.Stdw1Maint Reqd - Stud Weld 1 Maintenance Required FB2[252].29'; 8094 '~S001R10CN.I.Stdw1Reject - Stud Weld 1 art Reject Fault FB2[252].30'; 8095 '~S001R10CN.I.Rvt1Flt - Rivet Controller 1 Fault FB2[252].31'; 8096 '~S001R10CN.I.Rvt1DlyExcdd - Rivet Cntrl 1 Time Delay Exceeded Flt FB2[253].0'; 8097 '~S001R10CN.I.AutoPulledTipByp1 - Auto Pulled Tip Bypass 1 FB2[253].1'; 8098 '~S001R10CN.I.StdWld1EquipmentFlt - Stud Weld 1 Equipment Fault FB2[253].2'; 8099 '~S001R10CN.I.StdWld1BrcktNotPresent - Stud Weld 1 Bracket Not Pres FB2[253].3'; 8100 '~S001R10CN.I.PierceFlt - Pierce Fault FB2[253].4'; 8101 '~S001R10CN.I.NoVisionMeasErr - Vision System Measurement Error FB2[253].5'; 8102 '~S001R10CN.I.VisionSysCalErr - Vision System Calibration Fault FB2[253].6'; 8103 '~S001R10CN.I.VisionSysErr - Vision System Error FB2[253].7'; 8104 '~S001R10CN.I.RackOutOfTolerance - Vision Sys Rack Out Of Tolerance FB2[253].8'; 8105 '~S001R10CN.Ix.TorqFlt - Torque Not Ok FB2[253].9'; 8106 '~S001R10CN.Ix.MwFlt - Mig Weld Controller Fault FB2[253].10'; 8107 '~S001R10CN.Ix.MwWireStuckFlt - Mig Welder Wire Stuck FB2[253].11'; 8108 '~S001R10CN.Ix.MwWldFlt - Mig Welder Bad Bronze Weld Indicator Flt FB2[253].12'; 8109 '~S001R10CN.I.O.TipChngReqd1 - Weld Cntrl 1 Tip Change Required FB2[253].13'; 8110 '~S001R10CN.I.M.NutDetectFlt1 - Nut Welder 1 Nut Detection Fault FB2[253].14'; 8111 '~S001R10CN.I.M.NutProjFlt1 - Nut Welder 1 Weld Not In Tolerance FB2[253].15'; 8112 '~S001R10CN.M.WrongRivetAtNose - Remove Wrong Rivet At Nose FB2[253].16'; 8113 '~S001R10CN.Ix.MwWldLimitErr - Mig Welder CurrentVoltage Out of Tolerance FB2[253].17'; 8114 '~S001R10CN.Ix.MigRdy Mig Welder Not Ready FB2[253].18'; 8115 '~Spare FB2[253].19'; 8116 '~Spare FB2[253].20'; 8117 '~S001R10CN.I.Wc2WldFlt -Weld Controller 2 Weld Fault FB2[253].21'; 8118 '~S001R10CN.I.Wc2Flt - Weld Timer Flt - Depress Man Weld To Continue FB2[253].22'; 8119 '~S001R10CN.I.Wc2SGunFlt - Weld Controller 2 Servo Gun Fault FB2[253].23'; 8120 '~S001R10CN.I.Wc2SGunMtrTempFlt - Cntrl 2 Servo Gun Motor Over Temp FB2[253].24'; 8121 '~S001R10CN.I.Td2MtrFlt - Tip Dress 2 Motor Fault FB2[253].25'; 8122 '~S001R10CN.I.WC2XfmrTempFlt - Weld Cntrl 2 Transformer Over Temp FB2[253].26'; 8123 '~S001R10CN.I.AutoTipChng2Flt - Auto Tip Changer 2 Fault FB2[253].27'; 8124 '~S001R10CN.I.Slr2NotReady - Seal Controller 2 Not Ready FB2[253].28'; 8125 '~S001R10CN.I.Slr2MajorFlt - Seal Controller 2 Major Fault FB2[253].29'; 8126 '~S001R10CN.I.Slr2VolNotOk - Seal Controller 2 Volume Not Ok Fault FB2[253].30'; 8127 '~S001R10CN.I.Slr2PurgeFlt - Seal Controller 2 Purge Fault FB2[253].31'; 8128 '~S001R10CN.I.Slr2DoserNot Filled - Seal Cntrl 2 Doser Not Filled FB2[254].0'; 8129 '~S001R10CN.I.Slr2No2ClnMxr - Seal Cntrl2 No 2C In Mixer Fault FB2[254].1'; 8130 '~S001R10CN.I.Slr2NzlBroken - Seal Controller 2 Nozzle Broken Fault FB2[254].2'; 8131 '~S001R10CN.I.Slr2NozzleChgReq - Seal Cntrl2 Nozzle Change Reqd FB2[254].3'; 8132 '~S001R10CN.I.Slr2CycleInterrupted - Seal Cntrl2 Cycle Interrupted FB2[254].4'; 8133 '~S001R10CN.I.Stdw2Flt - Stud Weld 2 Weld Fault FB2[254].5'; 8134 '~S001R10CN.I.Stdw2DlyExcdd - Stud Weld 2 Time Delay Exceeded Flt FB2[254].6'; 8135 '~S001R10CN.I.Stdw2Maint Reqd - Stud Weld 2 Maintenance Required FB2[254].7'; 8136 '~S001R10CN.I.Stdw2Reject - Stud Weld 2 art Reject Fault FB2[254].8'; 8137 '~S001R10CN.I.Rvt2Flt - Rivet Controller 2 Fault FB2[254].9'; 8138 '~S001R10CN.I.Rvt2DlyExcdd - Rivet Cntrl 2 Time Delay Exceeded Flt FB2[254].10'; 8139 '~S001R10CN.I.AutoPulledTipByp2 - Auto Pulled Tip Bypass 2 FB2[254].11'; 8140 '~S001R10CN.I.StdWld2EquipmentFlt - Stud Weld 2 Equipment Fault FB2[254].12'; 8141 '~S001R10CN.I.StdWld2BrcktNotPresent - Stud Weld 2 Bracket Not Pres FB2[254].13'; 8142 '~S001R10CN.Ix.LsrWldMntrFlt - Seam Geometry/Laser Weld Monitor Flt FB2[254].14'; 8143 '~S001R10CN.Ix.LsrHeadFlt - Laser Head Fault FB2[254].15'; 8144 '~S001R10CN.Ix.LsrGlsFlt - Glass Fault FB2[254].16'; 8145 '~S001R10CN.Ix.LsrWhlFlt - Pressure Wheel Not In Range Fault FB2[254].17'; 8146 '~S001R10CN.Ix.LsrGeoFlt - Seam Geometry/Laser Bad Process Geo Flt FB2[254].18'; 8147 '~S001R10CN.Ix.LsrHdCollFlt - Laser Head Collision Fault FB2[254].19'; 8148 '~S001R10CN.Ix.LsrHdSysFlt - Laser Head System Fault FB2[254].20'; 8149 '~S001R10CN.Ix.LsrHdFar - Laser Head Far Fault FB2[254].21'; 8150 '~S001R10CN.Ix.LsrHdSftCollFlt - Laser Head Software Collision Flt FB2[254].22'; 8151 '~S001R10CN.I.O.TipChngReqd2 - Weld Cntrl 2 Tip Change Required FB2[254].23'; 8152 '~S001R10CN.I.M.NutDetectFlt2 - Nut Welder 2 Nut Detection Fault FB2[254].24'; 8153 '~S001R10CN.I.M.NutProjFlt2 - Nut Welder 2 Weld Not In Tolerance FB2[254].25'; 8154 '~S001R10CN.I.TCWrongToolInStand - Tool Changer Wrong Tool In Stand FB2[254].26'; 8155 '~Spare FB2[254].27'; 8156 '~Spare FB2[254].28'; 8157 '~Spare FB2[254].29'; 8158 '~Spare FB2[254].30'; 8159 '~Spare FB2[254].31'; 8160 '~S001R10CN.I.VisionCommOK - Vision System Comm Fault FB2[255].0'; 8161 '~S001R10CN.I.OutOfTolerance - Vision System Out Of Tolerance FB2[255].1'; 8162 '~S001R10CN.I.MeasureReject - Vision System Measure Reject FB2[255].2'; 8163 '~S001R10CN.I.VisionSysCalibrationFlt - Vision System Calibration Flt FB2[255].3'; 8164 '~S001R10CN.I.VisionSysFlt - Vision System Flt FB2[255].4'; 8165 '~Spare FB2[255].5'; 8166 '~Spare FB2[255].6'; 8167 '~Spare FB2[255].7'; 8168 '~Spare FB2[255].8'; 8169 '~Spare FB2[255].9'; 8170 '~Spare FB2[255].10'; 8171 '~Spare FB2[255].11'; 8172 '~Spare FB2[255].12'; 8173 '~Spare FB2[255].13'; 8174 '~Spare FB2[255].14'; 8175 '~Spare FB2[255].15'; 8176 '~Spare FB2[255].16'; 8177 '~Spare FB2[255].17'; 8178 '~S001R10CN.M.InteruptCyc - Laser Cyc Interupt Cut Wire And Reject Car FB2[255].18'; 8179 '~S001R10CN.M.SuspectPart Inspect Vehicle And Accept Or Reject FB2[255].19'; 8180 '~S001R10 Power Meter High Power Fault Detected FB2[255].20'; 8181 '~S001R10 Power Meter Low Power Fault Detected FB2[255].21'; 8182 '~Spare FB2[255].22'; 8183 '~Spare FB2[255].23'; 8184 '~Spare FB2[255].24'; 8185 '~Spare FB2[255].25'; 8186 '~Spare FB2[255].26'; 8187 '~Spare FB2[255].27'; 8188 '~Spare FB2[255].28'; 8189 '~Spare FB2[255].29'; 8190 '~Spare FB2[255].30'; 8191 '~Spare FB2[255].31'; 8192 '~Spare FB2[256].0'; 8193 '~Spare FB2[256].1'; 8194 '~Spare FB2[256].2'; 8195 '~Spare FB2[256].3'; 8196 '~Spare FB2[256].4'; 8197 '~Spare FB2[256].5'; 8198 '~Spare FB2[256].6'; 8199 '~Spare FB2[256].7'; 8200 '~Spare FB2[256].8'; 8201 '~Spare FB2[256].9'; 8202 '~Spare FB2[256].10'; 8203 '~Spare FB2[256].11'; 8204 '~Spare FB2[256].12'; 8205 '~Spare FB2[256].13'; 8206 '~Spare FB2[256].14'; 8207 '~Spare FB2[256].15'; 8208 '~Spare FB2[256].16'; 8209 '~Spare FB2[256].17'; 8210 '~Spare FB2[256].18'; 8211 '~Spare FB2[256].19'; 8212 '~Spare FB2[256].20'; 8213 '~Spare FB2[256].21'; 8214 '~Spare FB2[256].22'; 8215 '~Spare FB2[256].23'; 8216 '~Spare FB2[256].24'; 8217 '~Spare FB2[256].25'; 8218 '~Spare FB2[256].26'; 8219 '~Spare FB2[256].27'; 8220 '~Spare FB2[256].28'; 8221 '~Spare FB2[256].29'; 8222 '~Spare FB2[256].30'; 8223 '~Spare FB2[256].31'; 8224 '~Spare FB2[257].0'; 8225 '~Spare FB2[257].1'; 8226 '~Spare FB2[257].2'; 8227 '~Spare FB2[257].3'; 8228 '~Spare FB2[257].4'; 8229 '~Spare FB2[257].5'; 8230 '~Spare FB2[257].6'; 8231 '~Spare FB2[257].7'; 8232 '~Spare FB2[257].8'; 8233 '~Spare FB2[257].9'; 8234 '~Spare FB2[257].10'; 8235 '~Spare FB2[257].11'; 8236 '~Spare FB2[257].12'; 8237 '~Spare FB2[257].13'; 8238 '~Spare FB2[257].14'; 8239 '~Spare FB2[257].15'; 8240 '~Spare FB2[257].16'; 8241 '~Spare FB2[257].17'; 8242 '~Spare FB2[257].18'; 8243 '~Spare FB2[257].19'; 8244 '~Spare FB2[257].20'; 8245 '~Spare FB2[257].21'; 8246 '~Spare FB2[257].22'; 8247 '~Spare FB2[257].23'; 8248 '~Spare FB2[257].24'; 8249 '~Spare FB2[257].25'; 8250 '~Spare FB2[257].26'; 8251 '~Spare FB2[257].27'; 8252 '~Spare FB2[257].28'; 8253 '~Spare FB2[257].29'; 8254 '~Spare FB2[257].30'; 8255 '~Spare FB2[257].31'; 8256 '~Spare FB2[258].0'; 8257 '~Spare FB2[258].1'; 8258 '~Spare FB2[258].2'; 8259 '~Spare FB2[258].3'; 8260 '~Spare FB2[258].4'; 8261 '~Spare FB2[258].5'; 8262 '~Spare FB2[258].6'; 8263 '~Spare FB2[258].7'; 8264 '~Spare FB2[258].8'; 8265 '~Spare FB2[258].9'; 8266 '~Spare FB2[258].10'; 8267 '~Spare FB2[258].11'; 8268 '~Spare FB2[258].12'; 8269 '~Spare FB2[258].13'; 8270 '~Spare FB2[258].14'; 8271 '~Spare FB2[258].15'; 8272 '~Spare FB2[258].16'; 8273 '~Spare FB2[258].17'; 8274 '~Spare FB2[258].18'; 8275 '~Spare FB2[258].19'; 8276 '~Spare FB2[258].20'; 8277 '~Spare FB2[258].21'; 8278 '~Spare FB2[258].22'; 8279 '~Spare FB2[258].23'; 8280 '~Spare FB2[258].24'; 8281 '~Spare FB2[258].25'; 8282 '~Spare FB2[258].26'; 8283 '~Spare FB2[258].27'; 8284 '~Spare FB2[258].28'; 8285 '~Spare FB2[258].29'; 8286 '~Spare FB2[258].30'; 8287 '~Spare FB2[258].31'; 8288 '~Spare FB2[259].0'; 8289 '~Spare FB2[259].1'; 8290 '~Spare FB2[259].2'; 8291 '~Spare FB2[259].3'; 8292 '~Spare FB2[259].4'; 8293 '~Spare FB2[259].5'; 8294 '~Spare FB2[259].6'; 8295 '~Spare FB2[259].7'; 8296 '~Spare FB2[259].8'; 8297 '~Spare FB2[259].9'; 8298 '~Spare FB2[259].10'; 8299 '~Spare FB2[259].11'; 8300 '~Spare FB2[259].12'; 8301 '~Spare FB2[259].13'; 8302 '~Spare FB2[259].14'; 8303 '~Spare FB2[259].15'; 8304 '~Spare FB2[259].16'; 8305 '~Spare FB2[259].17'; 8306 '~Spare FB2[259].18'; 8307 '~Spare FB2[259].19'; 8308 '~Spare FB2[259].20'; 8309 '~Spare FB2[259].21'; 8310 '~Spare FB2[259].22'; 8311 '~Spare FB2[259].23'; 8312 '~Spare FB2[259].24'; 8313 '~Spare FB2[259].25'; 8314 '~Spare FB2[259].26'; 8315 '~Spare FB2[259].27'; 8316 '~Spare FB2[259].28'; 8317 '~Spare FB2[259].29'; 8318 '~Spare FB2[259].30'; 8319 '~Spare FB2[259].31'; 8320 '~S001R11CN.I.RbtCtrlFlt - Control Fault FB2[260].0'; 8321 '~S001R11CN.I.CollDetect - Collision Detect FB2[260].1'; 8322 '~S001R11CN.Ix.RbtPromptBox - View Prompt Box at Teach Pendant FB2[260].2'; 8323 '~Spare FB2[260].3'; 8324 '~Spare FB2[260].4'; 8325 '~Spare FB2[260].5'; 8326 '~Spare FB2[260].6'; 8327 '~Spare FB2[260].7'; 8328 '~Spare FB2[260].8'; 8329 '~Spare FB2[260].9'; 8330 '~Spare FB2[260].10'; 8331 '~S001R11CN.I.Wc1WldFlt -Weld Controller 1 Weld Fault FB2[260].11'; 8332 '~S001R11CN.I.Wc1Flt - Weld Timer Flt - Depress Man Weld To Continue FB2[260].12'; 8333 '~S001R11CN.I.Wc1SGunFlt - Weld Controller 1 Servo Gun Fault FB2[260].13'; 8334 '~S001R11CN.I.Wc1SGunMtrTempFlt - Cntrl 1 Servo Gun Motor Over Temp FB2[260].14'; 8335 '~S001R11CN.I.Td1MtrFlt - Tip Dress 1 Motor Fault FB2[260].15'; 8336 '~S001R11CN.I.WC1XfmrTempFlt - Weld Cntrl 1 Transformer Over Temp FB2[260].16'; 8337 '~S001R11CN.I.AutoTipChng1Flt - Auto Tip Changer 1 Fault FB2[260].17'; 8338 '~S001R11CN.I.Slr1NotReady - Seal Controller 1 Not Ready FB2[260].18'; 8339 '~S001R11CN.I.Slr1MajorFlt - Seal Controller 1 Major Fault FB2[260].19'; 8340 '~S001R11CN.I.Slr1VolNotOk - Seal 